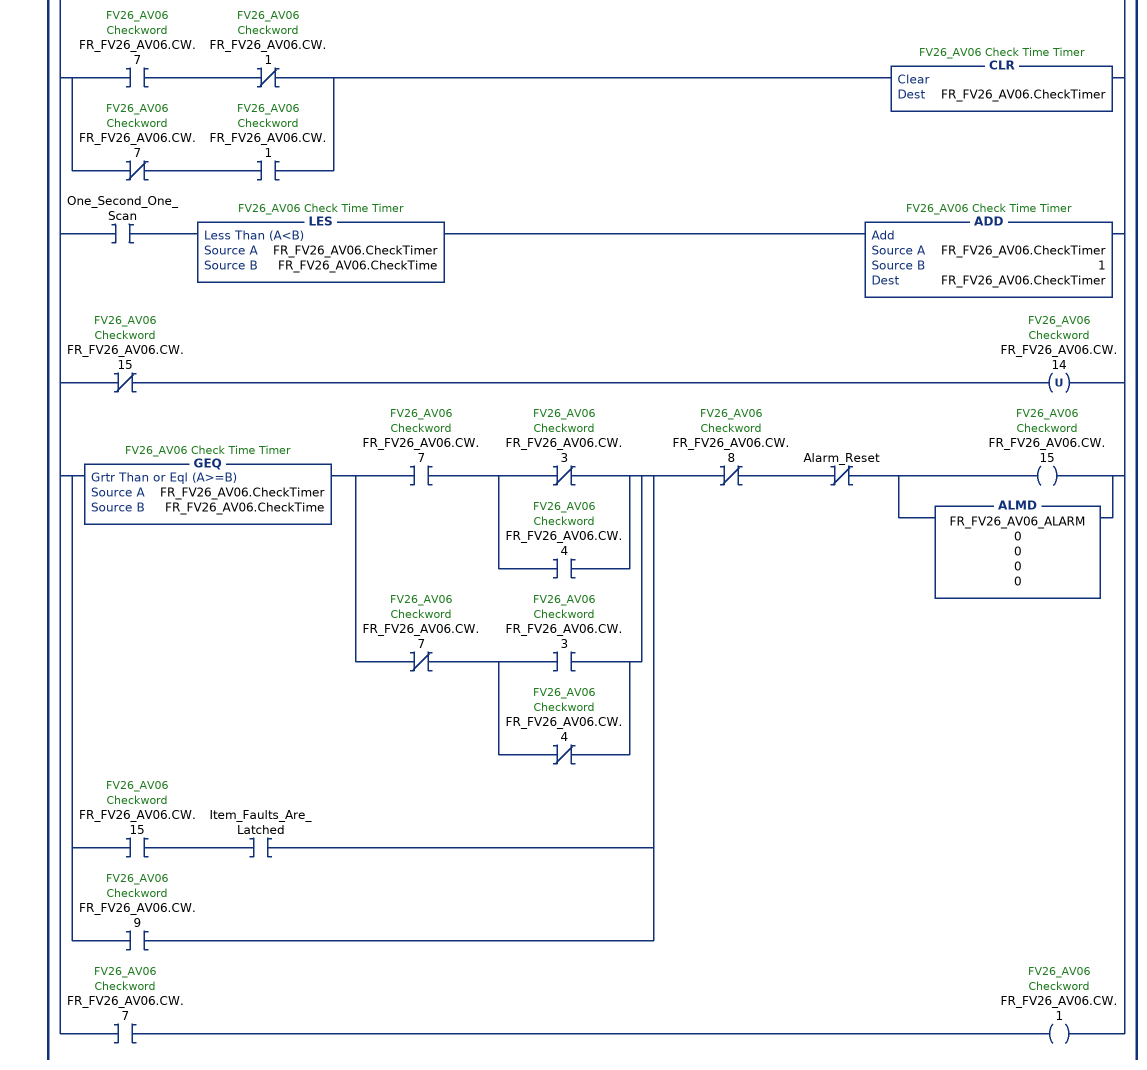
   4: [NEQ(FR_FV26_AV06.DriveBits,0) OTE(FR_FV26_AV06.CW.0) ,[XIC(FR_FV26_AV06.CW.0) XIO(FR_FV26_AV06.CW.6) ,XIC(FR_FV26_AV06.CW.5) XIC(FR_FV26_AV06.CW.6) ] OTE(FR_FV26_AV06.CW.7) ,XIC(FR_FV26_AV06.CW.7) OTE(FR_FV26_AV06_DR) ,XIC(S:FS) [OTU(FR_FV26_AV06.CW.6) ,LEQ(FR_FV26_AV06.CheckTime,0) MOV(Default_Check_Time,FR_FV26_AV06.CheckTime) ] ,[[XIC(FR_FV26_AV06_O) XIO(Item_Simulation_Flag) ,XIC(Item_Simulation_Flag) XIC(FR_FV26_AV06.CW.7) XIO(FR_FV26_AV06.CW.2) ] OTE(FR_FV26_AV06.CW.3) ,[XIC(FR_FV26_AV06_C) XIO(Item_Simulation_Flag) ,XIC(Item_Simulation_Flag) XIO(FR_FV26_AV06.CW.7) XIO(FR_FV26_AV06.CW.2) ] OTE(FR_FV26_AV06.CW.4) ] ,[XIC(FR_FV26_AV06.CW.7) XIO(FR_FV26_AV06.CW.1) ,XIO(FR_FV26_AV06.CW.7) XIC(FR_FV26_AV06.CW.1) ] CLR(FR_FV26_AV06.CheckTimer) ,XIC(One_Second_One_Scan) LES(FR_FV26_AV06.CheckTimer,FR_FV26_AV06.CheckTime) ADD(FR_FV26_AV06.CheckTimer,1,FR_FV26_AV06.CheckTimer) ,XIO(FR_FV26_AV06.CW.15) OTU(FR_FV26_AV06.CW.14) ,[GEQ(FR_FV26_AV06.CheckTimer,FR_FV26_AV06.CheckTime) [XIC(FR_FV26_AV06.CW.7) [XIO(FR_FV26_AV06.CW.3) ,XIC(FR_FV26_AV06.CW.4) ] ,XIO(FR_FV26_AV06.CW.7) [XIC(FR_FV26_AV06.CW.3) ,XIO(FR_FV26_AV06.CW.4) ] ] ,XIC(FR_FV26_AV06.CW.15) XIC(Item_Faults_Are_Latched) ,XIC(FR_FV26_AV06.CW.9) ] XIO(FR_FV26_AV06.CW.8) XIO(Alarm_Reset) [OTE(FR_FV26_AV06.CW.15) ,ALMD(FR_FV26_AV06_ALARM,0,0,0,0) ] ,XIC(FR_FV26_AV06.CW.7) OTE(FR_FV26_AV06.CW.1) ];
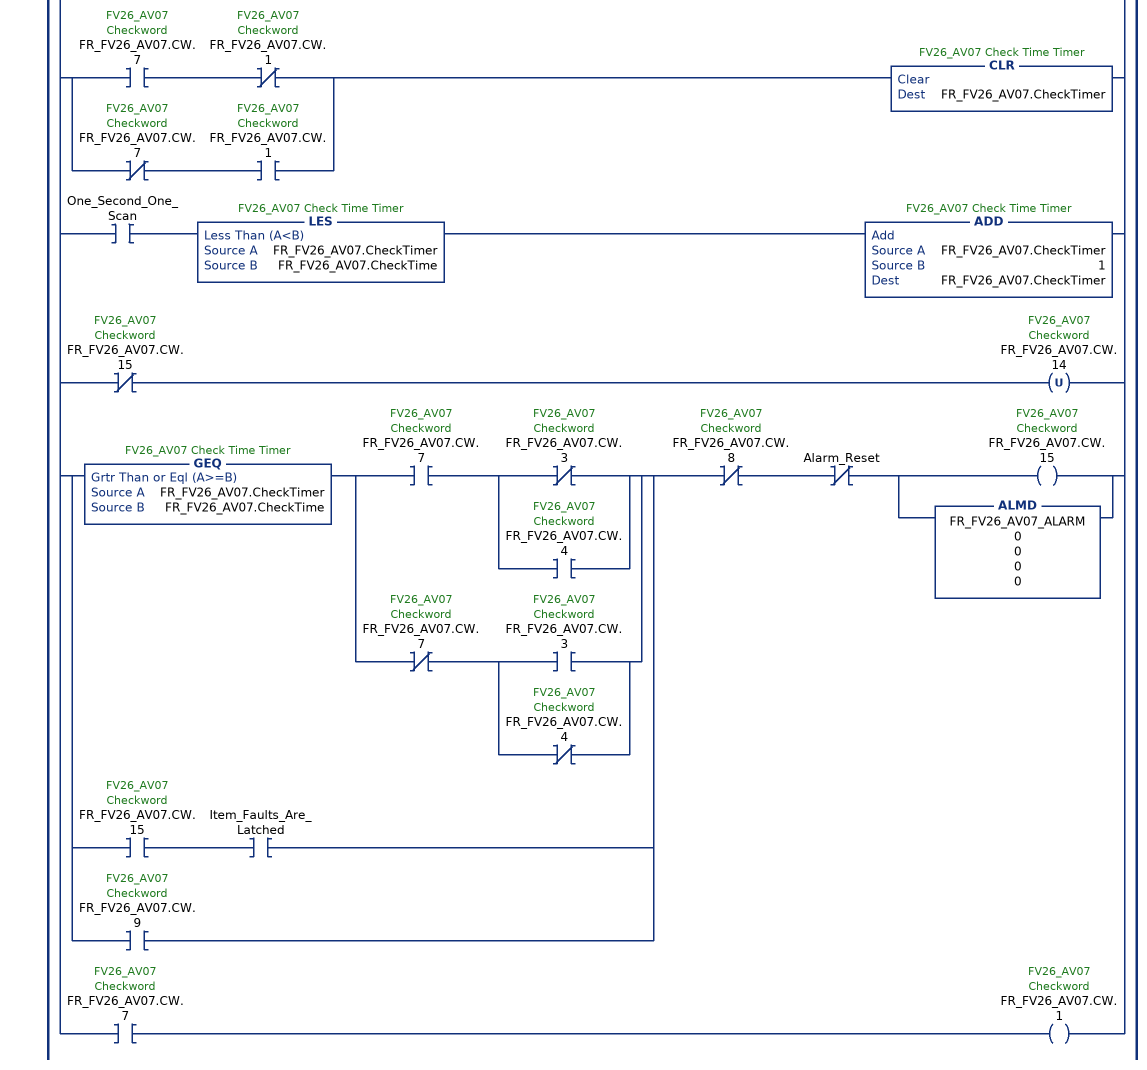
   5: [NEQ(FR_FV26_AV07.DriveBits,0) OTE(FR_FV26_AV07.CW.0) ,[XIC(FR_FV26_AV07.CW.0) XIO(FR_FV26_AV07.CW.6) ,XIC(FR_FV26_AV07.CW.5) XIC(FR_FV26_AV07.CW.6) ] OTE(FR_FV26_AV07.CW.7) ,XIC(FR_FV26_AV07.CW.7) OTE(FR_FV26_AV07_DR) ,XIC(S:FS) [OTU(FR_FV26_AV07.CW.6) ,LEQ(FR_FV26_AV07.CheckTime,0) MOV(Default_Check_Time,FR_FV26_AV07.CheckTime) ] ,[[XIC(FR_FV26_AV07_O) XIO(Item_Simulation_Flag) ,XIC(Item_Simulation_Flag) XIC(FR_FV26_AV07.CW.7) XIO(FR_FV26_AV07.CW.2) ] OTE(FR_FV26_AV07.CW.3) ,[XIC(FR_FV26_AV07_C) XIO(Item_Simulation_Flag) ,XIC(Item_Simulation_Flag) XIO(FR_FV26_AV07.CW.7) XIO(FR_FV26_AV07.CW.2) ] OTE(FR_FV26_AV07.CW.4) ] ,[XIC(FR_FV26_AV07.CW.7) XIO(FR_FV26_AV07.CW.1) ,XIO(FR_FV26_AV07.CW.7) XIC(FR_FV26_AV07.CW.1) ] CLR(FR_FV26_AV07.CheckTimer) ,XIC(One_Second_One_Scan) LES(FR_FV26_AV07.CheckTimer,FR_FV26_AV07.CheckTime) ADD(FR_FV26_AV07.CheckTimer,1,FR_FV26_AV07.CheckTimer) ,XIO(FR_FV26_AV07.CW.15) OTU(FR_FV26_AV07.CW.14) ,[GEQ(FR_FV26_AV07.CheckTimer,FR_FV26_AV07.CheckTime) [XIC(FR_FV26_AV07.CW.7) [XIO(FR_FV26_AV07.CW.3) ,XIC(FR_FV26_AV07.CW.4) ] ,XIO(FR_FV26_AV07.CW.7) [XIC(FR_FV26_AV07.CW.3) ,XIO(FR_FV26_AV07.CW.4) ] ] ,XIC(FR_FV26_AV07.CW.15) XIC(Item_Faults_Are_Latched) ,XIC(FR_FV26_AV07.CW.9) ] XIO(FR_FV26_AV07.CW.8) XIO(Alarm_Reset) [OTE(FR_FV26_AV07.CW.15) ,ALMD(FR_FV26_AV07_ALARM,0,0,0,0) ] ,XIC(FR_FV26_AV07.CW.7) OTE(FR_FV26_AV07.CW.1) ];
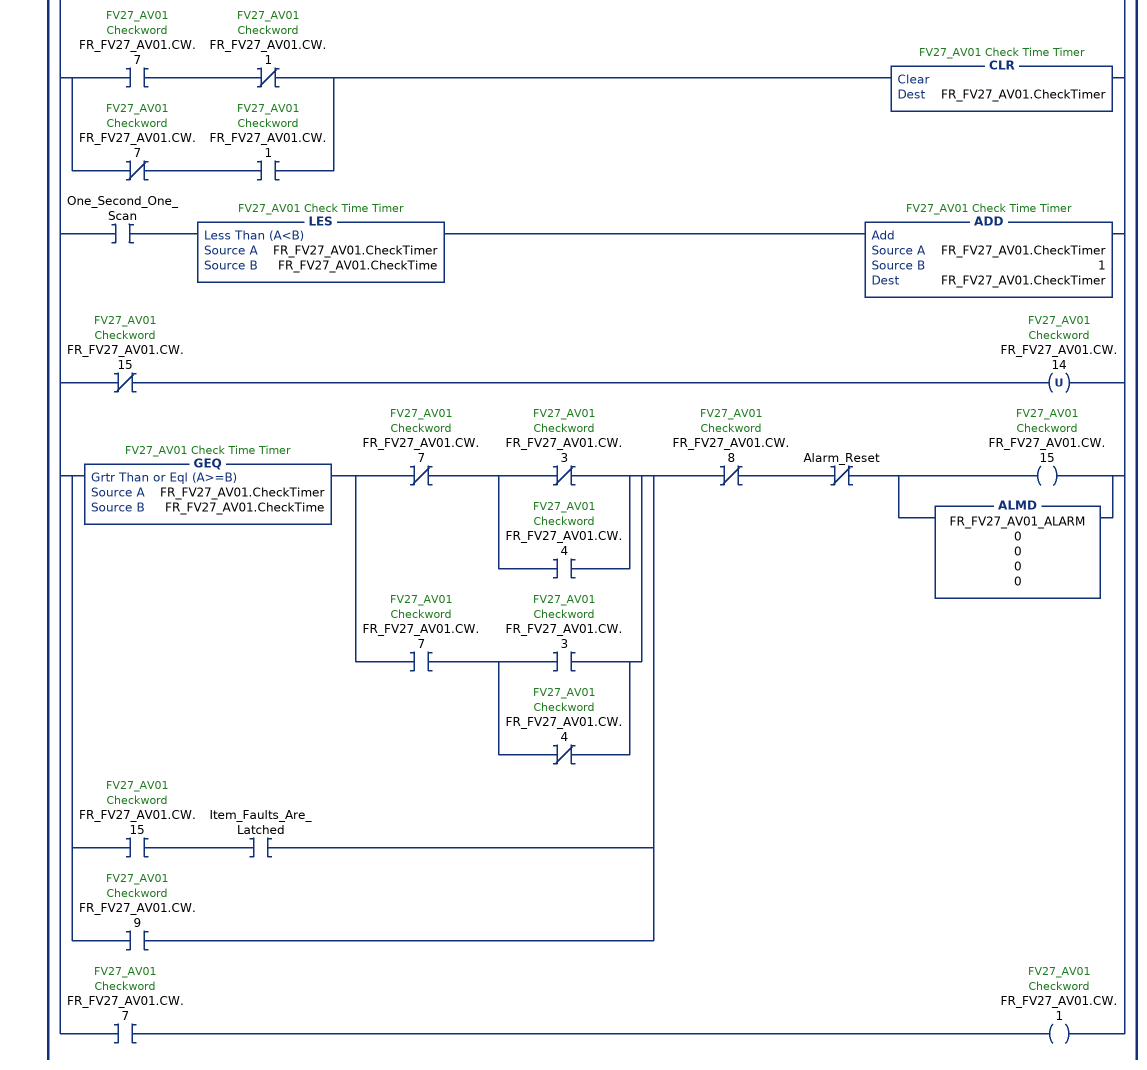
   6: [NEQ(FR_FV27_AV01.DriveBits,0) OTE(FR_FV27_AV01.CW.0) ,[XIC(FR_FV27_AV01.CW.0) XIO(FR_FV27_AV01.CW.6) ,XIC(FR_FV27_AV01.CW.5) XIC(FR_FV27_AV01.CW.6) ] OTE(FR_FV27_AV01.CW.7) ,XIC(FR_FV27_AV01.CW.7) OTE(FR_FV27_AV01_RDR) ,XIC(S:FS) [OTU(FR_FV27_AV01.CW.6) ,LEQ(FR_FV27_AV01.CheckTime,0) MOV(Default_Check_Time,FR_FV27_AV01.CheckTime) ] ,[[XIC(FR_FV27_AV01_C) XIO(Item_Simulation_Flag) ,XIC(Item_Simulation_Flag) XIO(FR_FV27_AV01.CW.7) XIO(FR_FV27_AV01.CW.2) ] OTE(FR_FV27_AV01.CW.3) ,[XIC(FR_FV27_AV01_O) XIO(Item_Simulation_Flag) ,XIC(Item_Simulation_Flag) XIC(FR_FV27_AV01.CW.7) XIO(FR_FV27_AV01.CW.2) ] OTE(FR_FV27_AV01.CW.4) ] ,[XIC(FR_FV27_AV01.CW.7) XIO(FR_FV27_AV01.CW.1) ,XIO(FR_FV27_AV01.CW.7) XIC(FR_FV27_AV01.CW.1) ] CLR(FR_FV27_AV01.CheckTimer) ,XIC(One_Second_One_Scan) LES(FR_FV27_AV01.CheckTimer,FR_FV27_AV01.CheckTime) ADD(FR_FV27_AV01.CheckTimer,1,FR_FV27_AV01.CheckTimer) ,XIO(FR_FV27_AV01.CW.15) OTU(FR_FV27_AV01.CW.14) ,[GEQ(FR_FV27_AV01.CheckTimer,FR_FV27_AV01.CheckTime) [XIO(FR_FV27_AV01.CW.7) [XIO(FR_FV27_AV01.CW.3) ,XIC(FR_FV27_AV01.CW.4) ] ,XIC(FR_FV27_AV01.CW.7) [XIC(FR_FV27_AV01.CW.3) ,XIO(FR_FV27_AV01.CW.4) ] ] ,XIC(FR_FV27_AV01.CW.15) XIC(Item_Faults_Are_Latched) ,XIC(FR_FV27_AV01.CW.9) ] XIO(FR_FV27_AV01.CW.8) XIO(Alarm_Reset) [OTE(FR_FV27_AV01.CW.15) ,ALMD(FR_FV27_AV01_ALARM,0,0,0,0) ] ,XIC(FR_FV27_AV01.CW.7) OTE(FR_FV27_AV01.CW.1) ];
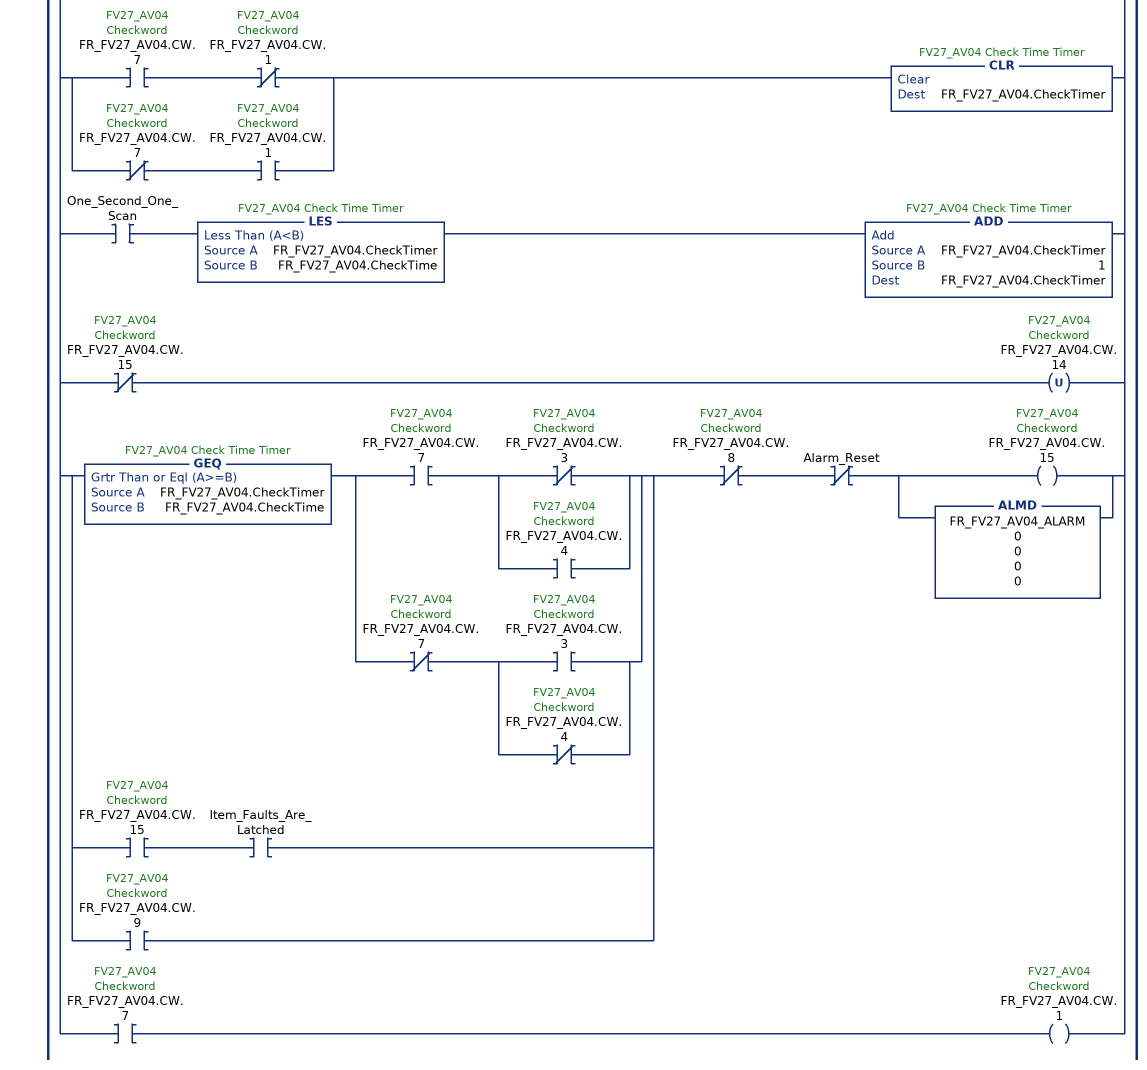
   7: [NEQ(FR_FV27_AV04.DriveBits,0) OTE(FR_FV27_AV04.CW.0) ,[XIC(FR_FV27_AV04.CW.0) XIO(FR_FV27_AV04.CW.6) ,XIC(FR_FV27_AV04.CW.5) XIC(FR_FV27_AV04.CW.6) ] OTE(FR_FV27_AV04.CW.7) ,XIC(FR_FV27_AV04.CW.7) OTE(FR_FV27_AV04_DR) ,XIC(S:FS) [OTU(FR_FV27_AV04.CW.6) ,LEQ(FR_FV27_AV04.CheckTime,0) MOV(Default_Check_Time,FR_FV27_AV04.CheckTime) ] ,[[XIC(FR_FV27_AV04_O) XIO(Item_Simulation_Flag) ,XIC(Item_Simulation_Flag) XIC(FR_FV27_AV04.CW.7) XIO(FR_FV27_AV04.CW.2) ] OTE(FR_FV27_AV04.CW.3) ,[XIC(FR_FV27_AV04_C) XIO(Item_Simulation_Flag) ,XIC(Item_Simulation_Flag) XIO(FR_FV27_AV04.CW.7) XIO(FR_FV27_AV04.CW.2) ] OTE(FR_FV27_AV04.CW.4) ] ,[XIC(FR_FV27_AV04.CW.7) XIO(FR_FV27_AV04.CW.1) ,XIO(FR_FV27_AV04.CW.7) XIC(FR_FV27_AV04.CW.1) ] CLR(FR_FV27_AV04.CheckTimer) ,XIC(One_Second_One_Scan) LES(FR_FV27_AV04.CheckTimer,FR_FV27_AV04.CheckTime) ADD(FR_FV27_AV04.CheckTimer,1,FR_FV27_AV04.CheckTimer) ,XIO(FR_FV27_AV04.CW.15) OTU(FR_FV27_AV04.CW.14) ,[GEQ(FR_FV27_AV04.CheckTimer,FR_FV27_AV04.CheckTime) [XIC(FR_FV27_AV04.CW.7) [XIO(FR_FV27_AV04.CW.3) ,XIC(FR_FV27_AV04.CW.4) ] ,XIO(FR_FV27_AV04.CW.7) [XIC(FR_FV27_AV04.CW.3) ,XIO(FR_FV27_AV04.CW.4) ] ] ,XIC(FR_FV27_AV04.CW.15) XIC(Item_Faults_Are_Latched) ,XIC(FR_FV27_AV04.CW.9) ] XIO(FR_FV27_AV04.CW.8) XIO(Alarm_Reset) [OTE(FR_FV27_AV04.CW.15) ,ALMD(FR_FV27_AV04_ALARM,0,0,0,0) ] ,XIC(FR_FV27_AV04.CW.7) OTE(FR_FV27_AV04.CW.1) ];
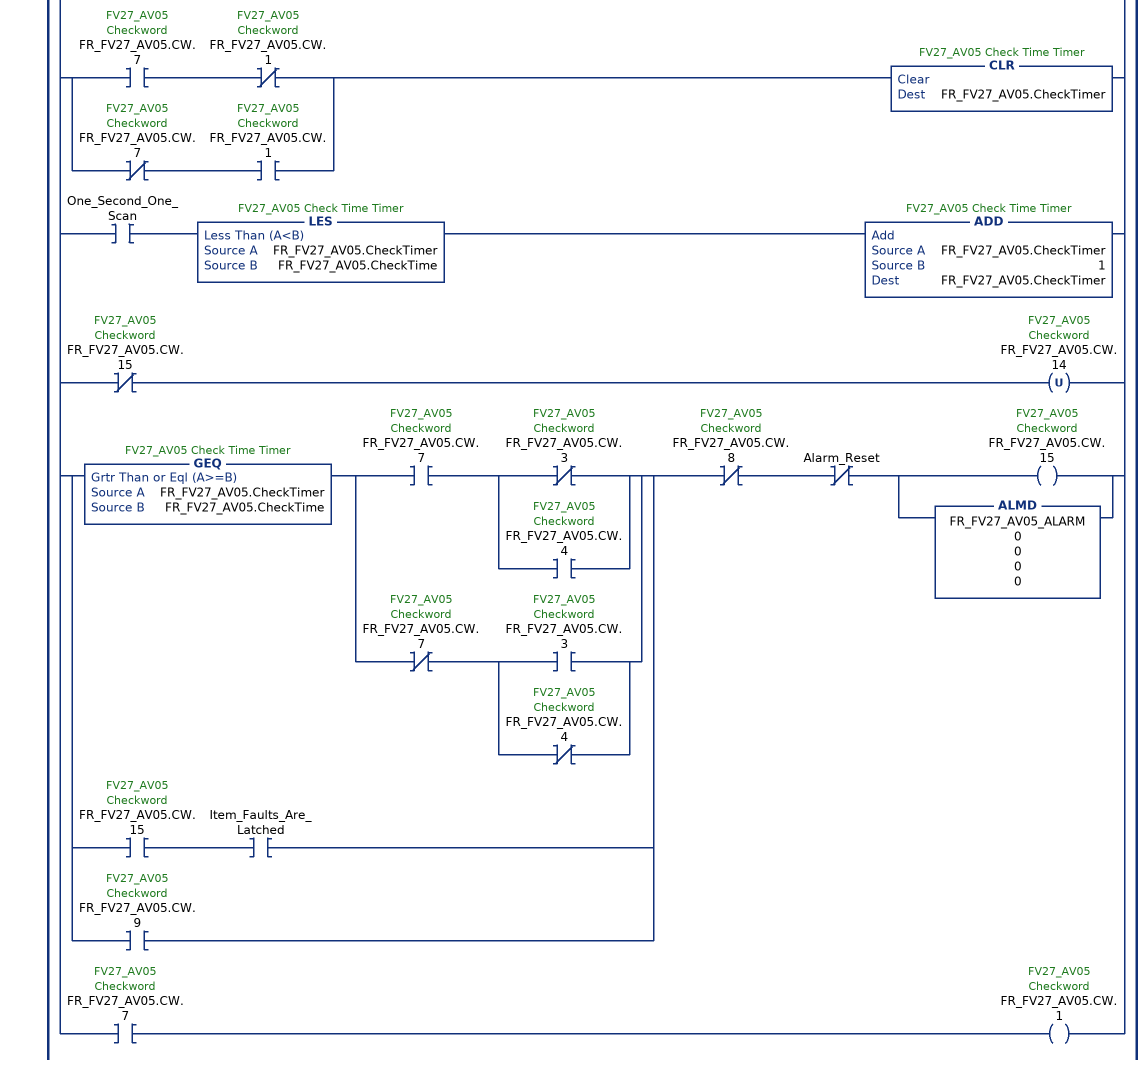
   8: [NEQ(FR_FV27_AV05.DriveBits,0) OTE(FR_FV27_AV05.CW.0) ,[XIC(FR_FV27_AV05.CW.0) XIO(FR_FV27_AV05.CW.6) ,XIC(FR_FV27_AV05.CW.5) XIC(FR_FV27_AV05.CW.6) ] OTE(FR_FV27_AV05.CW.7) ,XIC(FR_FV27_AV05.CW.7) OTE(FR_FV27_AV05_DR) ,XIC(S:FS) [OTU(FR_FV27_AV05.CW.6) ,LEQ(FR_FV27_AV05.CheckTime,0) MOV(Default_Check_Time,FR_FV27_AV05.CheckTime) ] ,[[XIC(FR_FV27_AV05_O) XIO(Item_Simulation_Flag) ,XIC(Item_Simulation_Flag) XIC(FR_FV27_AV05.CW.7) XIO(FR_FV27_AV05.CW.2) ] OTE(FR_FV27_AV05.CW.3) ,[XIC(FR_FV27_AV05_C) XIO(Item_Simulation_Flag) ,XIC(Item_Simulation_Flag) XIO(FR_FV27_AV05.CW.7) XIO(FR_FV27_AV05.CW.2) ] OTE(FR_FV27_AV05.CW.4) ] ,[XIC(FR_FV27_AV05.CW.7) XIO(FR_FV27_AV05.CW.1) ,XIO(FR_FV27_AV05.CW.7) XIC(FR_FV27_AV05.CW.1) ] CLR(FR_FV27_AV05.CheckTimer) ,XIC(One_Second_One_Scan) LES(FR_FV27_AV05.CheckTimer,FR_FV27_AV05.CheckTime) ADD(FR_FV27_AV05.CheckTimer,1,FR_FV27_AV05.CheckTimer) ,XIO(FR_FV27_AV05.CW.15) OTU(FR_FV27_AV05.CW.14) ,[GEQ(FR_FV27_AV05.CheckTimer,FR_FV27_AV05.CheckTime) [XIC(FR_FV27_AV05.CW.7) [XIO(FR_FV27_AV05.CW.3) ,XIC(FR_FV27_AV05.CW.4) ] ,XIO(FR_FV27_AV05.CW.7) [XIC(FR_FV27_AV05.CW.3) ,XIO(FR_FV27_AV05.CW.4) ] ] ,XIC(FR_FV27_AV05.CW.15) XIC(Item_Faults_Are_Latched) ,XIC(FR_FV27_AV05.CW.9) ] XIO(FR_FV27_AV05.CW.8) XIO(Alarm_Reset) [OTE(FR_FV27_AV05.CW.15) ,ALMD(FR_FV27_AV05_ALARM,0,0,0,0) ] ,XIC(FR_FV27_AV05.CW.7) OTE(FR_FV27_AV05.CW.1) ];
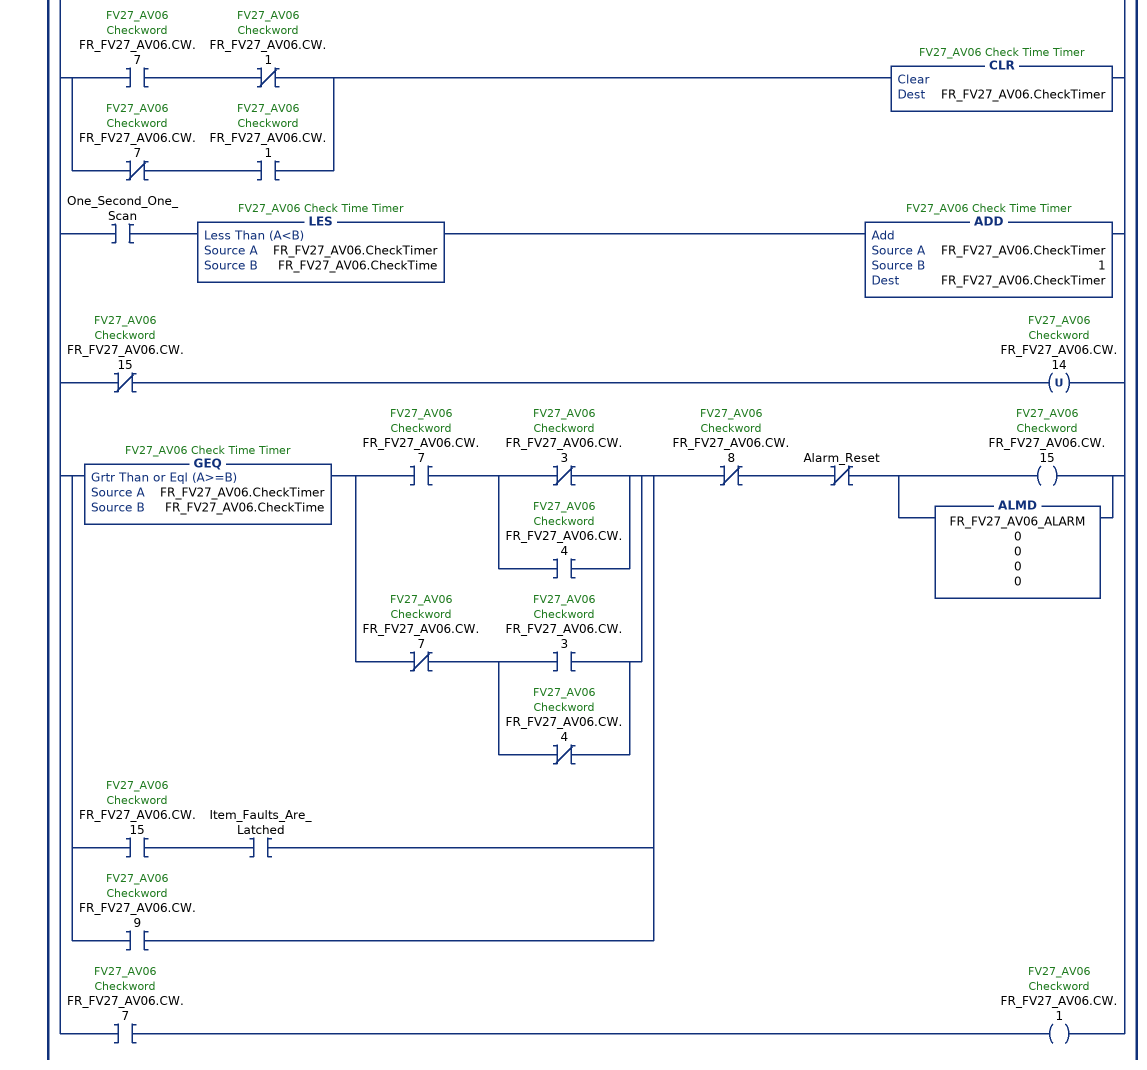
   9: [NEQ(FR_FV27_AV06.DriveBits,0) OTE(FR_FV27_AV06.CW.0) ,[XIC(FR_FV27_AV06.CW.0) XIO(FR_FV27_AV06.CW.6) ,XIC(FR_FV27_AV06.CW.5) XIC(FR_FV27_AV06.CW.6) ] OTE(FR_FV27_AV06.CW.7) ,XIC(FR_FV27_AV06.CW.7) OTE(FR_FV27_AV06_DR) ,XIC(S:FS) [OTU(FR_FV27_AV06.CW.6) ,LEQ(FR_FV27_AV06.CheckTime,0) MOV(Default_Check_Time,FR_FV27_AV06.CheckTime) ] ,[[XIC(FR_FV27_AV06_O) XIO(Item_Simulation_Flag) ,XIC(Item_Simulation_Flag) XIC(FR_FV27_AV06.CW.7) XIO(FR_FV27_AV06.CW.2) ] OTE(FR_FV27_AV06.CW.3) ,[XIC(FR_FV27_AV06_C) XIO(Item_Simulation_Flag) ,XIC(Item_Simulation_Flag) XIO(FR_FV27_AV06.CW.7) XIO(FR_FV27_AV06.CW.2) ] OTE(FR_FV27_AV06.CW.4) ] ,[XIC(FR_FV27_AV06.CW.7) XIO(FR_FV27_AV06.CW.1) ,XIO(FR_FV27_AV06.CW.7) XIC(FR_FV27_AV06.CW.1) ] CLR(FR_FV27_AV06.CheckTimer) ,XIC(One_Second_One_Scan) LES(FR_FV27_AV06.CheckTimer,FR_FV27_AV06.CheckTime) ADD(FR_FV27_AV06.CheckTimer,1,FR_FV27_AV06.CheckTimer) ,XIO(FR_FV27_AV06.CW.15) OTU(FR_FV27_AV06.CW.14) ,[GEQ(FR_FV27_AV06.CheckTimer,FR_FV27_AV06.CheckTime) [XIC(FR_FV27_AV06.CW.7) [XIO(FR_FV27_AV06.CW.3) ,XIC(FR_FV27_AV06.CW.4) ] ,XIO(FR_FV27_AV06.CW.7) [XIC(FR_FV27_AV06.CW.3) ,XIO(FR_FV27_AV06.CW.4) ] ] ,XIC(FR_FV27_AV06.CW.15) XIC(Item_Faults_Are_Latched) ,XIC(FR_FV27_AV06.CW.9) ] XIO(FR_FV27_AV06.CW.8) XIO(Alarm_Reset) [OTE(FR_FV27_AV06.CW.15) ,ALMD(FR_FV27_AV06_ALARM,0,0,0,0) ] ,XIC(FR_FV27_AV06.CW.7) OTE(FR_FV27_AV06.CW.1) ];
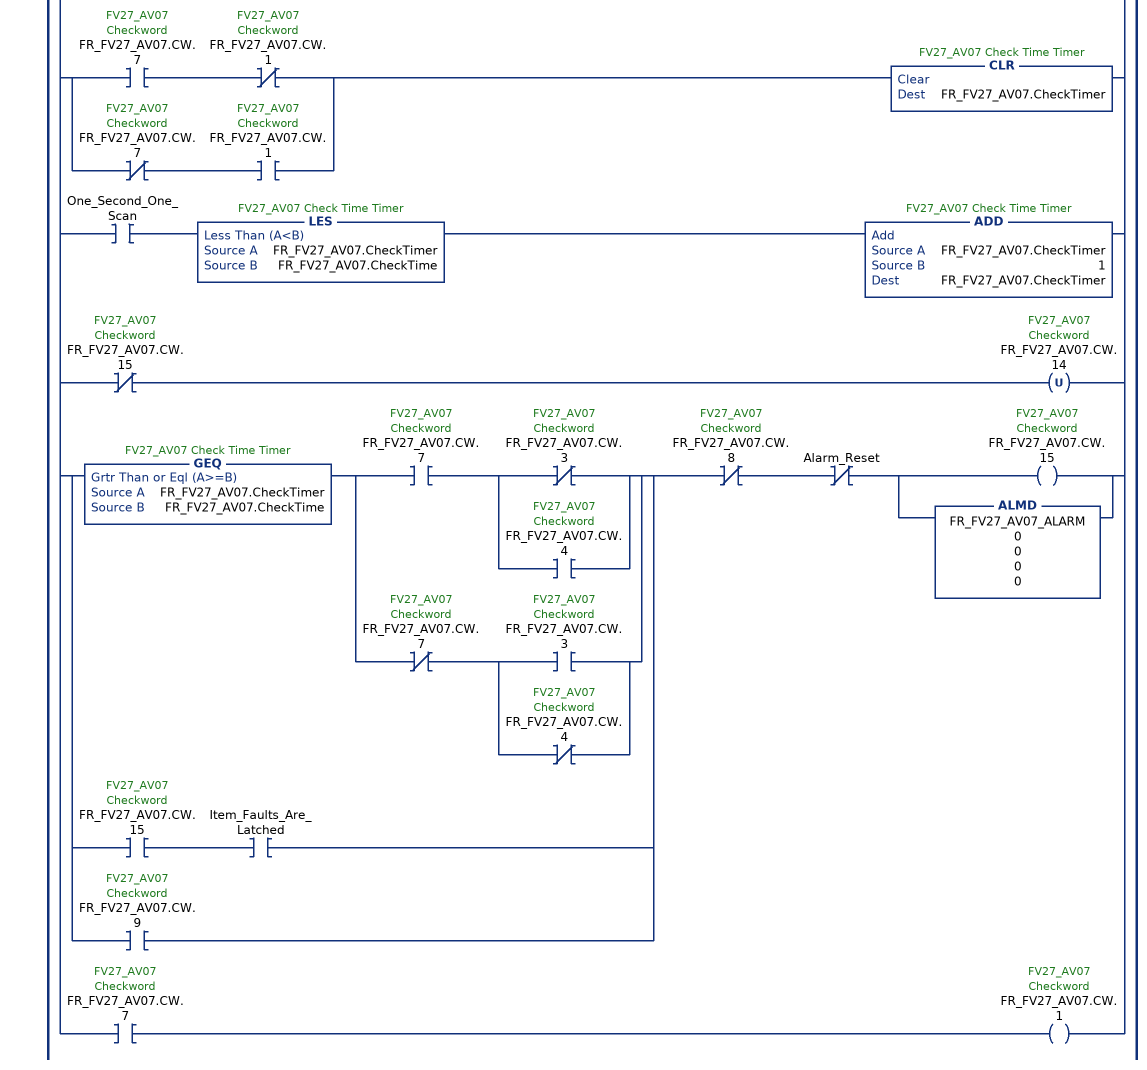
   10: [NEQ(FR_FV27_AV07.DriveBits,0) OTE(FR_FV27_AV07.CW.0) ,[XIC(FR_FV27_AV07.CW.0) XIO(FR_FV27_AV07.CW.6) ,XIC(FR_FV27_AV07.CW.5) XIC(FR_FV27_AV07.CW.6) ] OTE(FR_FV27_AV07.CW.7) ,XIC(FR_FV27_AV07.CW.7) OTE(FR_FV27_AV07_DR) ,XIC(S:FS) [OTU(FR_FV27_AV07.CW.6) ,LEQ(FR_FV27_AV07.CheckTime,0) MOV(Default_Check_Time,FR_FV27_AV07.CheckTime) ] ,[[XIC(FR_FV27_AV07_O) XIO(Item_Simulation_Flag) ,XIC(Item_Simulation_Flag) XIC(FR_FV27_AV07.CW.7) XIO(FR_FV27_AV07.CW.2) ] OTE(FR_FV27_AV07.CW.3) ,[XIC(FR_FV27_AV07_C) XIO(Item_Simulation_Flag) ,XIC(Item_Simulation_Flag) XIO(FR_FV27_AV07.CW.7) XIO(FR_FV27_AV07.CW.2) ] OTE(FR_FV27_AV07.CW.4) ] ,[XIC(FR_FV27_AV07.CW.7) XIO(FR_FV27_AV07.CW.1) ,XIO(FR_FV27_AV07.CW.7) XIC(FR_FV27_AV07.CW.1) ] CLR(FR_FV27_AV07.CheckTimer) ,XIC(One_Second_One_Scan) LES(FR_FV27_AV07.CheckTimer,FR_FV27_AV07.CheckTime) ADD(FR_FV27_AV07.CheckTimer,1,FR_FV27_AV07.CheckTimer) ,XIO(FR_FV27_AV07.CW.15) OTU(FR_FV27_AV07.CW.14) ,[GEQ(FR_FV27_AV07.CheckTimer,FR_FV27_AV07.CheckTime) [XIC(FR_FV27_AV07.CW.7) [XIO(FR_FV27_AV07.CW.3) ,XIC(FR_FV27_AV07.CW.4) ] ,XIO(FR_FV27_AV07.CW.7) [XIC(FR_FV27_AV07.CW.3) ,XIO(FR_FV27_AV07.CW.4) ] ] ,XIC(FR_FV27_AV07.CW.15) XIC(Item_Faults_Are_Latched) ,XIC(FR_FV27_AV07.CW.9) ] XIO(FR_FV27_AV07.CW.8) XIO(Alarm_Reset) [OTE(FR_FV27_AV07.CW.15) ,ALMD(FR_FV27_AV07_ALARM,0,0,0,0) ] ,XIC(FR_FV27_AV07.CW.7) OTE(FR_FV27_AV07.CW.1) ];
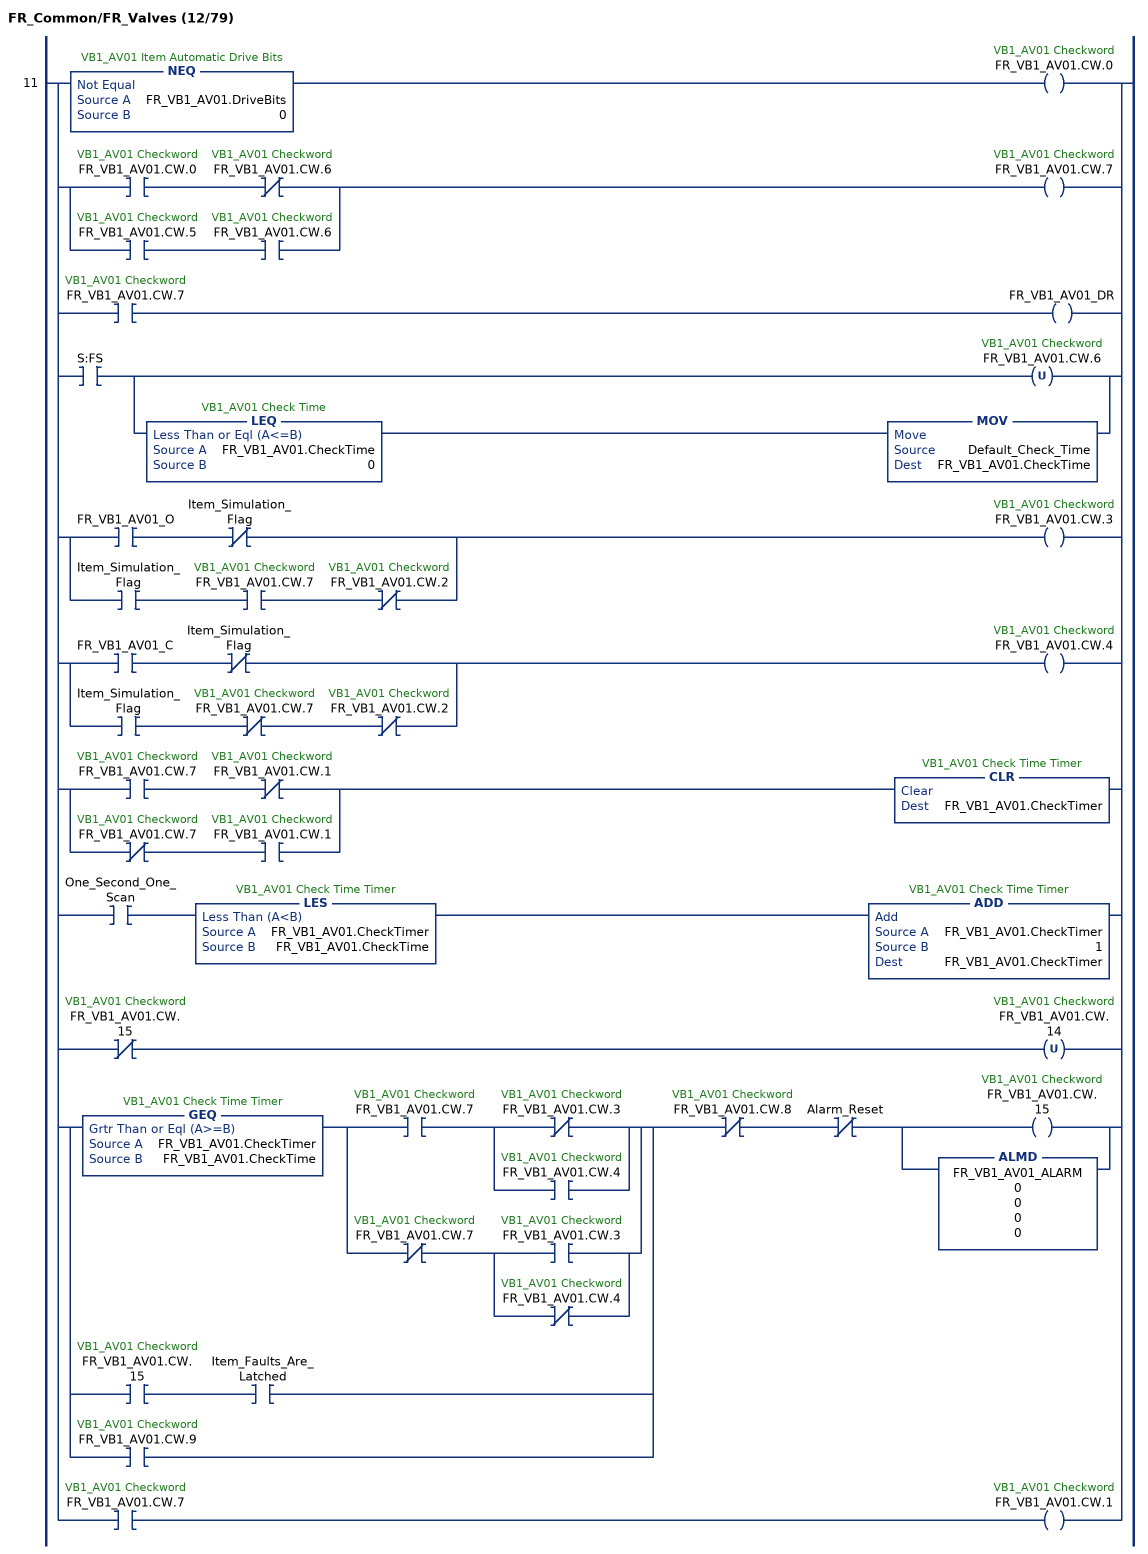
   11: [NEQ(FR_VB1_AV01.DriveBits,0) OTE(FR_VB1_AV01.CW.0) ,[XIC(FR_VB1_AV01.CW.0) XIO(FR_VB1_AV01.CW.6) ,XIC(FR_VB1_AV01.CW.5) XIC(FR_VB1_AV01.CW.6) ] OTE(FR_VB1_AV01.CW.7) ,XIC(FR_VB1_AV01.CW.7) OTE(FR_VB1_AV01_DR) ,XIC(S:FS) [OTU(FR_VB1_AV01.CW.6) ,LEQ(FR_VB1_AV01.CheckTime,0) MOV(Default_Check_Time,FR_VB1_AV01.CheckTime) ] ,[[XIC(FR_VB1_AV01_O) XIO(Item_Simulation_Flag) ,XIC(Item_Simulation_Flag) XIC(FR_VB1_AV01.CW.7) XIO(FR_VB1_AV01.CW.2) ] OTE(FR_VB1_AV01.CW.3) ,[XIC(FR_VB1_AV01_C) XIO(Item_Simulation_Flag) ,XIC(Item_Simulation_Flag) XIO(FR_VB1_AV01.CW.7) XIO(FR_VB1_AV01.CW.2) ] OTE(FR_VB1_AV01.CW.4) ] ,[XIC(FR_VB1_AV01.CW.7) XIO(FR_VB1_AV01.CW.1) ,XIO(FR_VB1_AV01.CW.7) XIC(FR_VB1_AV01.CW.1) ] CLR(FR_VB1_AV01.CheckTimer) ,XIC(One_Second_One_Scan) LES(FR_VB1_AV01.CheckTimer,FR_VB1_AV01.CheckTime) ADD(FR_VB1_AV01.CheckTimer,1,FR_VB1_AV01.CheckTimer) ,XIO(FR_VB1_AV01.CW.15) OTU(FR_VB1_AV01.CW.14) ,[GEQ(FR_VB1_AV01.CheckTimer,FR_VB1_AV01.CheckTime) [XIC(FR_VB1_AV01.CW.7) [XIO(FR_VB1_AV01.CW.3) ,XIC(FR_VB1_AV01.CW.4) ] ,XIO(FR_VB1_AV01.CW.7) [XIC(FR_VB1_AV01.CW.3) ,XIO(FR_VB1_AV01.CW.4) ] ] ,XIC(FR_VB1_AV01.CW.15) XIC(Item_Faults_Are_Latched) ,XIC(FR_VB1_AV01.CW.9) ] XIO(FR_VB1_AV01.CW.8) XIO(Alarm_Reset) [OTE(FR_VB1_AV01.CW.15) ,ALMD(FR_VB1_AV01_ALARM,0,0,0,0) ] ,XIC(FR_VB1_AV01.CW.7) OTE(FR_VB1_AV01.CW.1) ];
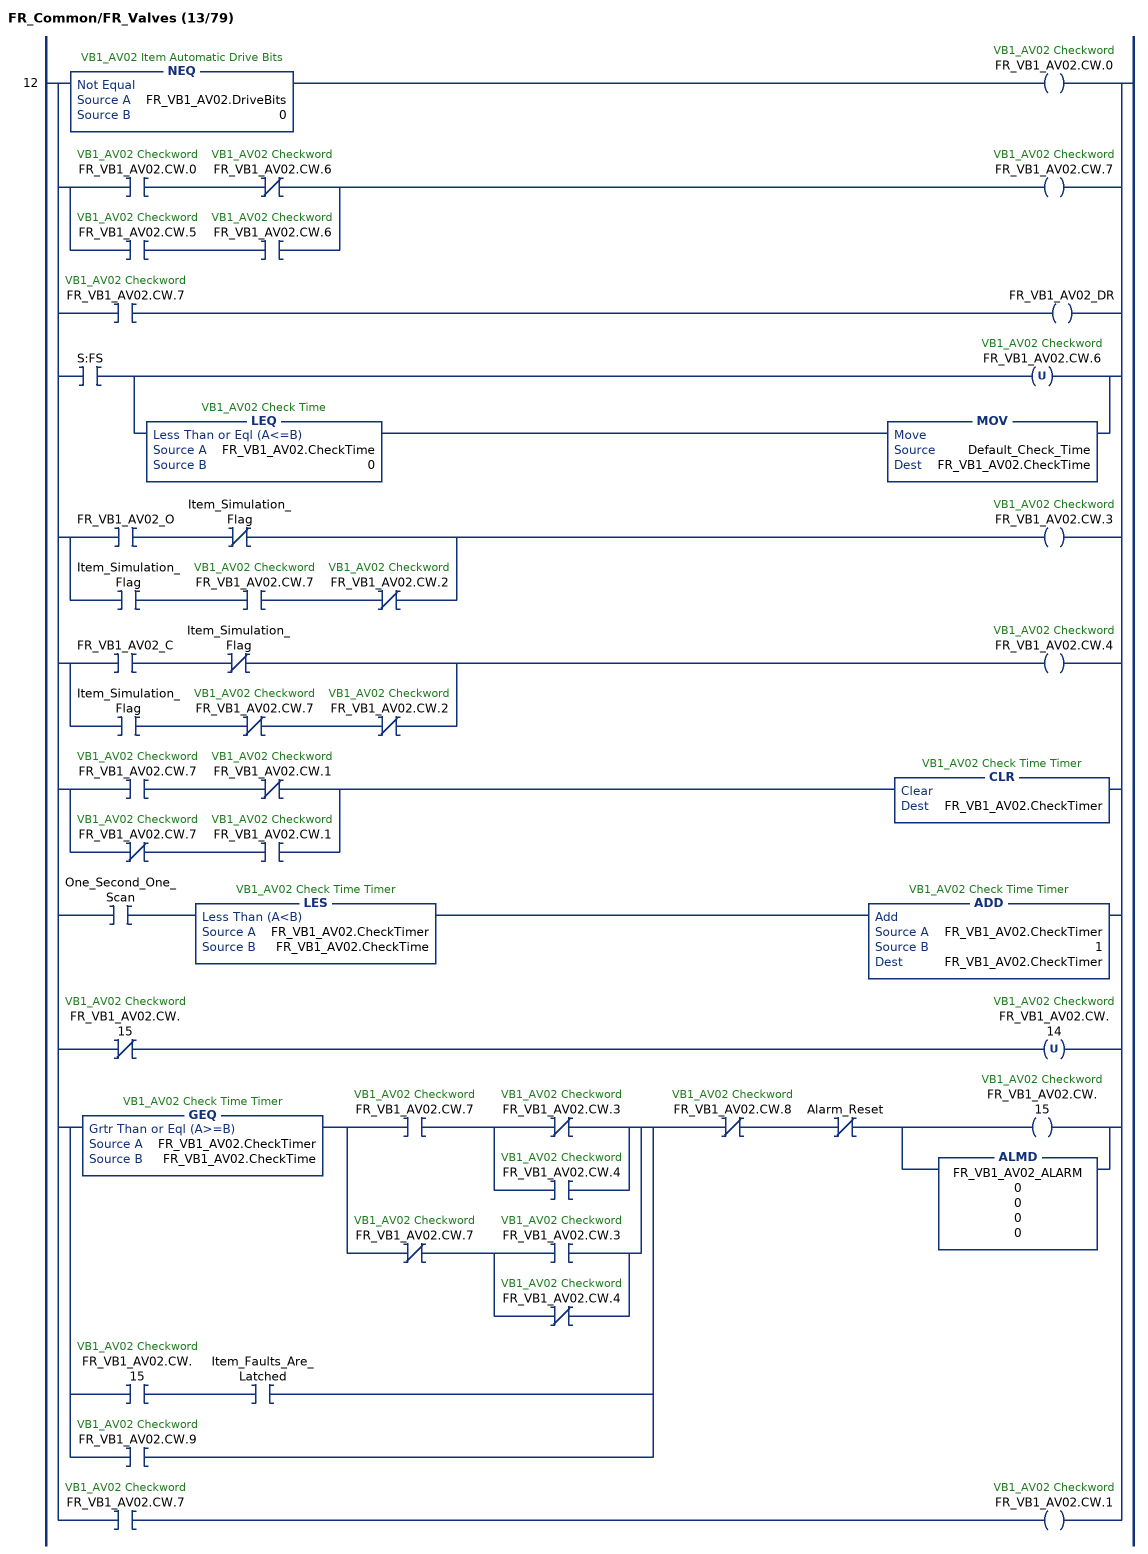
   12: [NEQ(FR_VB1_AV02.DriveBits,0) OTE(FR_VB1_AV02.CW.0) ,[XIC(FR_VB1_AV02.CW.0) XIO(FR_VB1_AV02.CW.6) ,XIC(FR_VB1_AV02.CW.5) XIC(FR_VB1_AV02.CW.6) ] OTE(FR_VB1_AV02.CW.7) ,XIC(FR_VB1_AV02.CW.7) OTE(FR_VB1_AV02_DR) ,XIC(S:FS) [OTU(FR_VB1_AV02.CW.6) ,LEQ(FR_VB1_AV02.CheckTime,0) MOV(Default_Check_Time,FR_VB1_AV02.CheckTime) ] ,[[XIC(FR_VB1_AV02_O) XIO(Item_Simulation_Flag) ,XIC(Item_Simulation_Flag) XIC(FR_VB1_AV02.CW.7) XIO(FR_VB1_AV02.CW.2) ] OTE(FR_VB1_AV02.CW.3) ,[XIC(FR_VB1_AV02_C) XIO(Item_Simulation_Flag) ,XIC(Item_Simulation_Flag) XIO(FR_VB1_AV02.CW.7) XIO(FR_VB1_AV02.CW.2) ] OTE(FR_VB1_AV02.CW.4) ] ,[XIC(FR_VB1_AV02.CW.7) XIO(FR_VB1_AV02.CW.1) ,XIO(FR_VB1_AV02.CW.7) XIC(FR_VB1_AV02.CW.1) ] CLR(FR_VB1_AV02.CheckTimer) ,XIC(One_Second_One_Scan) LES(FR_VB1_AV02.CheckTimer,FR_VB1_AV02.CheckTime) ADD(FR_VB1_AV02.CheckTimer,1,FR_VB1_AV02.CheckTimer) ,XIO(FR_VB1_AV02.CW.15) OTU(FR_VB1_AV02.CW.14) ,[GEQ(FR_VB1_AV02.CheckTimer,FR_VB1_AV02.CheckTime) [XIC(FR_VB1_AV02.CW.7) [XIO(FR_VB1_AV02.CW.3) ,XIC(FR_VB1_AV02.CW.4) ] ,XIO(FR_VB1_AV02.CW.7) [XIC(FR_VB1_AV02.CW.3) ,XIO(FR_VB1_AV02.CW.4) ] ] ,XIC(FR_VB1_AV02.CW.15) XIC(Item_Faults_Are_Latched) ,XIC(FR_VB1_AV02.CW.9) ] XIO(FR_VB1_AV02.CW.8) XIO(Alarm_Reset) [OTE(FR_VB1_AV02.CW.15) ,ALMD(FR_VB1_AV02_ALARM,0,0,0,0) ] ,XIC(FR_VB1_AV02.CW.7) OTE(FR_VB1_AV02.CW.1) ];
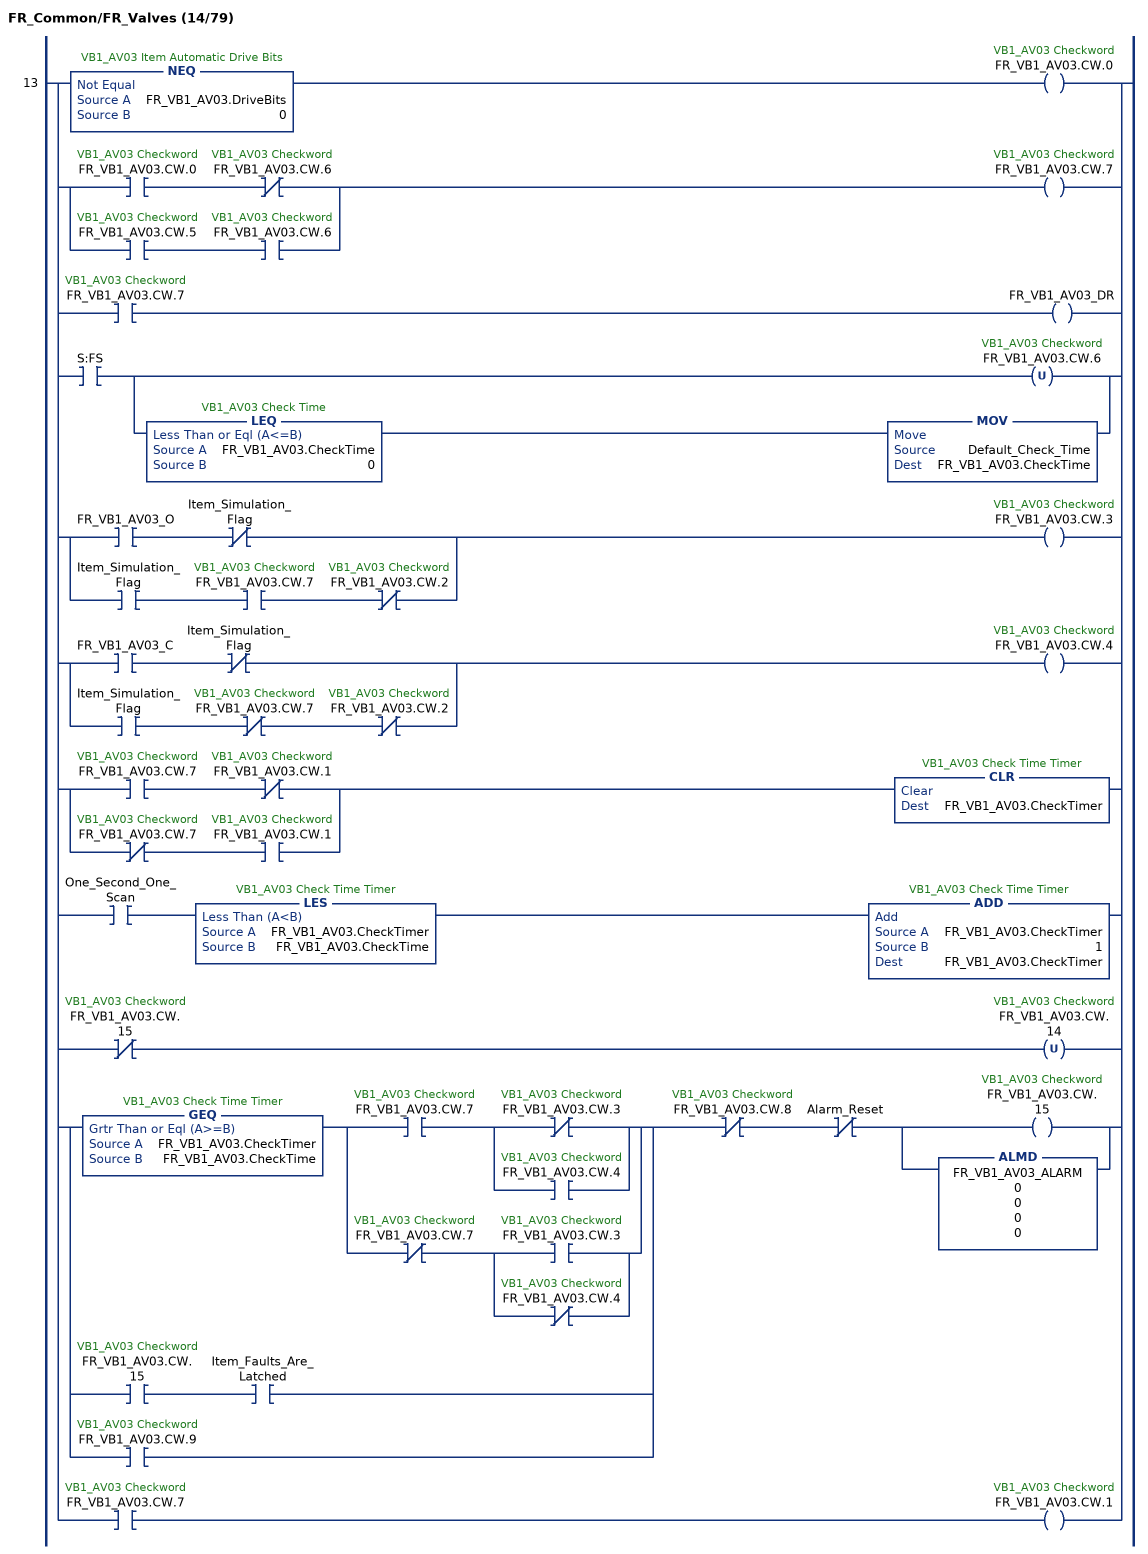
   13: [NEQ(FR_VB1_AV03.DriveBits,0) OTE(FR_VB1_AV03.CW.0) ,[XIC(FR_VB1_AV03.CW.0) XIO(FR_VB1_AV03.CW.6) ,XIC(FR_VB1_AV03.CW.5) XIC(FR_VB1_AV03.CW.6) ] OTE(FR_VB1_AV03.CW.7) ,XIC(FR_VB1_AV03.CW.7) OTE(FR_VB1_AV03_DR) ,XIC(S:FS) [OTU(FR_VB1_AV03.CW.6) ,LEQ(FR_VB1_AV03.CheckTime,0) MOV(Default_Check_Time,FR_VB1_AV03.CheckTime) ] ,[[XIC(FR_VB1_AV03_O) XIO(Item_Simulation_Flag) ,XIC(Item_Simulation_Flag) XIC(FR_VB1_AV03.CW.7) XIO(FR_VB1_AV03.CW.2) ] OTE(FR_VB1_AV03.CW.3) ,[XIC(FR_VB1_AV03_C) XIO(Item_Simulation_Flag) ,XIC(Item_Simulation_Flag) XIO(FR_VB1_AV03.CW.7) XIO(FR_VB1_AV03.CW.2) ] OTE(FR_VB1_AV03.CW.4) ] ,[XIC(FR_VB1_AV03.CW.7) XIO(FR_VB1_AV03.CW.1) ,XIO(FR_VB1_AV03.CW.7) XIC(FR_VB1_AV03.CW.1) ] CLR(FR_VB1_AV03.CheckTimer) ,XIC(One_Second_One_Scan) LES(FR_VB1_AV03.CheckTimer,FR_VB1_AV03.CheckTime) ADD(FR_VB1_AV03.CheckTimer,1,FR_VB1_AV03.CheckTimer) ,XIO(FR_VB1_AV03.CW.15) OTU(FR_VB1_AV03.CW.14) ,[GEQ(FR_VB1_AV03.CheckTimer,FR_VB1_AV03.CheckTime) [XIC(FR_VB1_AV03.CW.7) [XIO(FR_VB1_AV03.CW.3) ,XIC(FR_VB1_AV03.CW.4) ] ,XIO(FR_VB1_AV03.CW.7) [XIC(FR_VB1_AV03.CW.3) ,XIO(FR_VB1_AV03.CW.4) ] ] ,XIC(FR_VB1_AV03.CW.15) XIC(Item_Faults_Are_Latched) ,XIC(FR_VB1_AV03.CW.9) ] XIO(FR_VB1_AV03.CW.8) XIO(Alarm_Reset) [OTE(FR_VB1_AV03.CW.15) ,ALMD(FR_VB1_AV03_ALARM,0,0,0,0) ] ,XIC(FR_VB1_AV03.CW.7) OTE(FR_VB1_AV03.CW.1) ];
